(* Logix 5000 project; controller _GigaDiscovery vendor 1 type 14 code 244 rev 35.11; software revision 35.03; part 14 of 23 *)
(* tags used below, declared in another part *)
   Timer : TIMER[60];
   All_Rack_Closed_Mem : BOOL;
   Automatic_E_Stop_Cl_0 : DINT;
   Automatic_E_Stop_Cl_1 : DINT;
   DC_Field_Motor_7 : UDT_CROUT;   // DC Field Motor 7 Gondola Contactor -Q16101E -Q16103E
   DC_Field_Pylon_Motors : UDT_CROUT;   // DC Field Pylon Motors Contactor -Q10101E -Q10103E
   Emergencies_CL0 : DINT[8];
   Emergencies_CL1 : DINT[14];
   FeedBack_Drives_Contactors : BOOL;
   Gondola_Drive_Enable : UDT_CROUT;   // Gondola Drive Ch1-Ch2 Start Enable Contactors -Q16105E -Q16107E
   I_Compressor_Min_Pressure : BOOL;   // Line Pressure Switch - Minimum Pressure -S21504B
   I_EStop_Pb_OCC1 : UDT_DCI_STOP_TEST;   // +OCC E-stop -S30301F
   I_EStop_Pb_OCC2 : UDT_DCI_STOP_TEST;   // +OCC2 E-Stop -S28502F
   I_Gate_ENTER_G01_Closed : UDT_DCM;   // GATE ENTER (G01) -B25204I
   I_Gate_EXIT_G05_Closed : UDT_DCM;   // GATE EXIT (G05) -B25304I
   I_Gate_OPERATOR_Closed : UDT_DCM;   // GATE 4 OPERATOR RFID SENSOR - MOP -B25404J
   I_Gates_Closed : UDT_DCM;   // Gate Closed RFID series -B24802J
   I_OCC1_Stop_Cycle_PB : BOOL;   // Stop Cycle -S30308F
   I_OCC2_ACONFIRM : BOOL;   // OCC2 Allow Main CONFIRM -S28602F
   I_OCC2_Disable : UDT_DCM;   // OCC 2 CONTROL DISABLE Page 310
   I_OCC2_Stop_Cycle_PB : BOOL;   // Stop Cycle -S28606F
   I_OCC_LockOut_Motion : UDT_DCM;   // OCC -Lockout Motion -Q31203E
   I_OCC_Memory_Footpedal : BOOL;
   I_OCC_Operator_Enable_Key : BOOL;   // OCC Console Enabled -S30305F
   I_Operator_Footpedal : BOOL;   // Operator Footpedal -S30901F
   I_Platform_Line_Min_Pressure_Switch : BOOL;   // Platform Line Minimum Pressure Switch -S21511B
   I_Platform_Line_Unlock_Pressure_Switch : BOOL;   // Unlock Platform Line Pressure Switch -S22006B
   I_Platform_Opened : UDT_DCM;   // Platform Opened RFID Series -Q23801J -Q23807J
   I_RESTRAINTS_MainValve_Cosed : BOOL;   // Main Valve Close Limit Switch -B40508I
   I_RESTRAINTS_PressureswitchCompressor : BOOL;   // RESTRAINTS Main Valve Pressure Switch -S40602J
   I_Start_PB : Start_AOI;   // Primary console Strat Push botton Right and Left -S30401F -S30403F
   Mem_All_Rack_Sensor_OFF : BOOL;
   Mem_RESTRAINTS_closed_Correctly : BOOL;
   No_Automatic_E_Stop_Cl_0_Request : BOOL;
   No_Automatic_E_Stop_Cl_1_Request : BOOL;
   No_Emergencies_CL0 : BOOL;
   No_Emergencies_CL1 : BOOL;
   No_Sfty : Std_to_Sfty;
   O_Platform_MainValve : UDT_CROUT;   // Platform main valve B21902I
   O_RESTRAINTS_MainValve : UDT_CROUT;   // Main Valve -B40501I
   Pb_Platform_Stop : BOOL;   // Platform Stop Command -S30608F
   Platform_Open_Cycle : Sequencer;
   Platform_Open_Permissive : Permissive;
   PltaformOpeneded_CycleComplete : BOOL;   // Rilevazione Piattaforme aperte con ciclo Completato
   Power_On_Delay : BOOL;
   ProofTest_Req : BOOL;
   Pylon_Contactor_OFF : BOOL;
   Pylon_Start_Drive_1_2 : UDT_CROUT;   // Pylon Start Drive 1 - 2 Contactors -Q9002H -Q9004H -Q10202G
   Pylon_Start_Drive_3_4 : UDT_CROUT;   // Pylon Start Drive 3 - 4 Contactors -Q9005H -Q9007H -Q12202G
   Pylon_Start_Drive_5_6 : UDT_CROUT;   // Pylon Start Drive 5 - 6 Contactors -Q9009E -Q9011E4 -Q14202G -Q14202G
   Pylon_Stopped_At_Home : BOOL;   // 5s
   Reset_Pulse : BOOL;
   RESTRAINTS_ChA_Open_Memory : BOOL;
   RESTRAINTS_ChB_Open_Memory : BOOL;
   RESTRAINTS_Closed : BOOL;   // All RESTRAINTS Closed
   RESTRAINTS_Rack_Sector_ON : BOOL;
   RESTRAINTS_Sector_Enable_OFF : BOOL;   // ALL RESTRAINTS rack commands OFF
   RESTRAINTS_Unlock_Valve_Pressure : BOOL;
   Start_Permissive : Permissive;
   Start_Permissive2 : Permissive;
   Start_Platform_AutoCycle_Pylon : BOOL;
   Start_Stop_Cycle : Sequencer;
   Start_TOF : TIMER;
   Valve_Proof_Test_Ok : BOOL;
(* S_Alarms, continued *)

ROUTINE _08_Gates   (* ladder *)
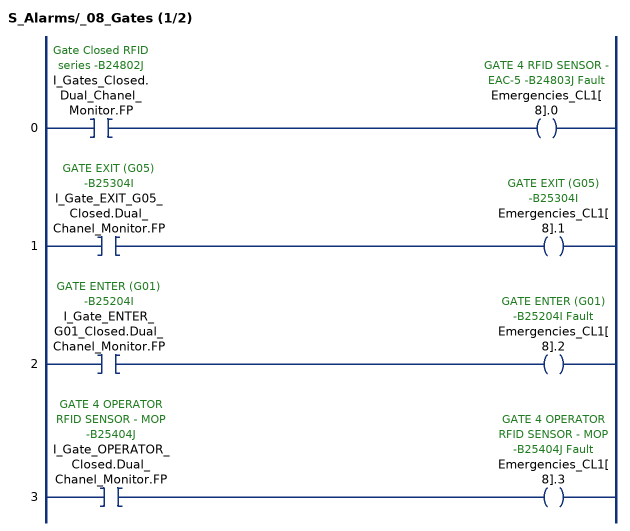
   0: XIC(I_Gates_Closed.Dual_Chanel_Monitor.FP)OTE(Emergencies_CL1[8].0);
   1: XIC(I_Gate_EXIT_G05_Closed.Dual_Chanel_Monitor.FP)OTE(Emergencies_CL1[8].1);
   2: XIC(I_Gate_ENTER_G01_Closed.Dual_Chanel_Monitor.FP)OTE(Emergencies_CL1[8].2);
   3: XIC(I_Gate_OPERATOR_Closed.Dual_Chanel_Monitor.FP)OTE(Emergencies_CL1[8].3);
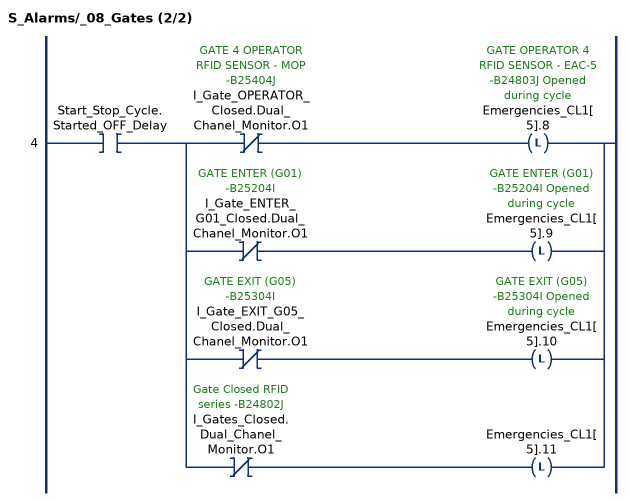
   4: XIC(Start_Stop_Cycle.Started_OFF_Delay)[XIO(I_Gate_OPERATOR_Closed.Dual_Chanel_Monitor.O1) OTL(Emergencies_CL1[5].8) ,XIO(I_Gate_ENTER_G01_Closed.Dual_Chanel_Monitor.O1) OTL(Emergencies_CL1[5].9) ,XIO(I_Gate_EXIT_G05_Closed.Dual_Chanel_Monitor.O1) OTL(Emergencies_CL1[5].10) ,XIO(I_Gates_Closed.Dual_Chanel_Monitor.O1) OTL(Emergencies_CL1[5].11) ];
END_ROUTINE

ROUTINE Main   (* ladder *)
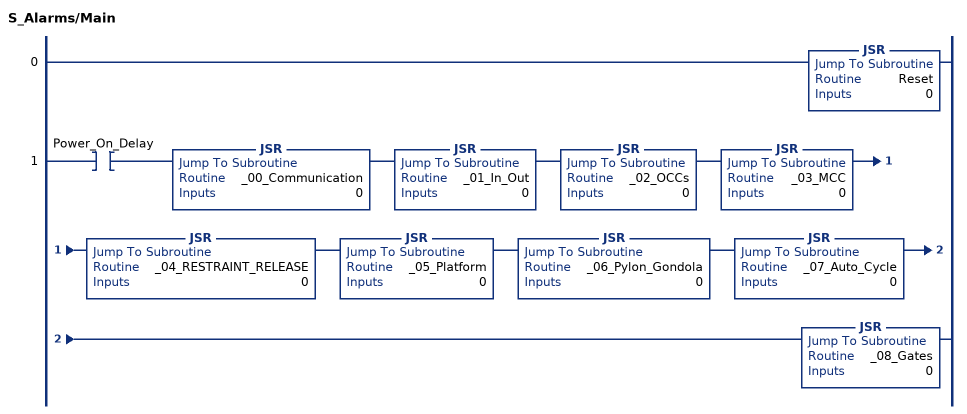
   0: JSR(Reset,0);
   1: XIC(Power_On_Delay)JSR(_00_Communication,0)JSR(_01_In_Out,0)JSR(_02_OCCs,0)JSR(_03_MCC,0)JSR(_04_RESTRAINT_RELEASE,0)JSR(_05_Platform,0)JSR(_06_Pylon_Gondola,0)JSR(_07_Auto_Cycle,0)JSR(_08_Gates,0);
END_ROUTINE

ROUTINE Reset   (* ladder *)
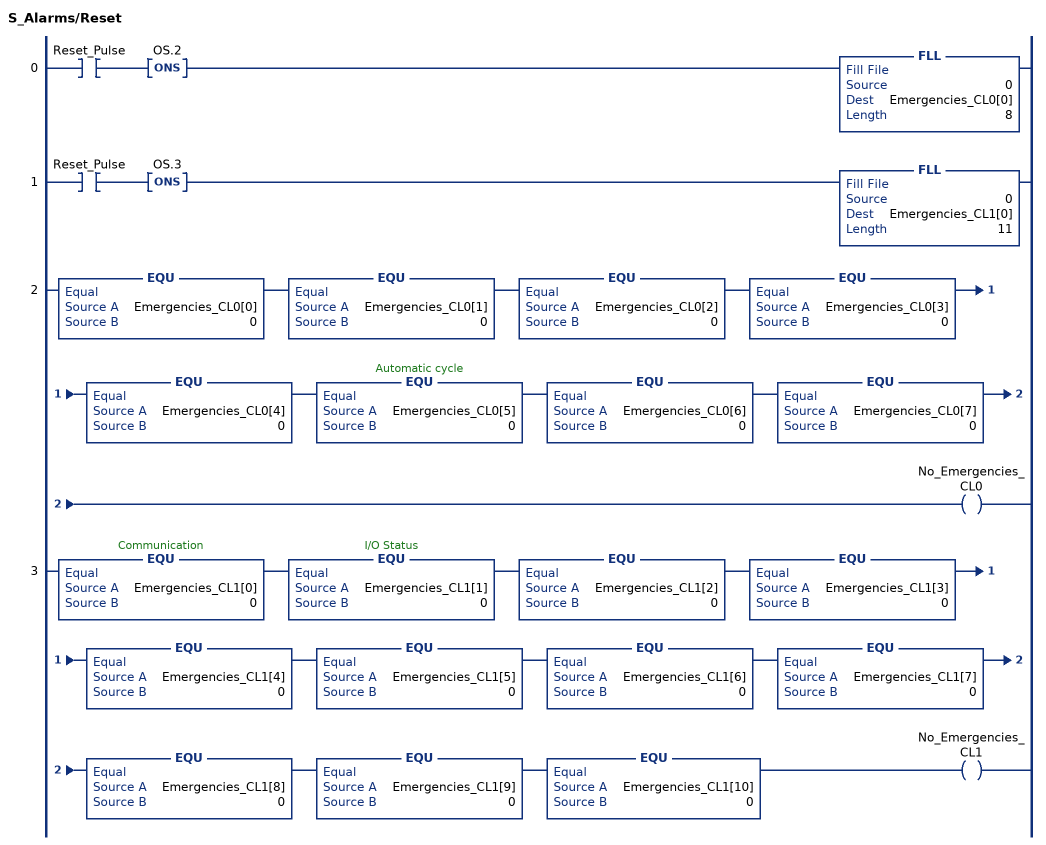
   0: XIC(Reset_Pulse)ONS(OS.2)FLL(0,Emergencies_CL0[0],8);
   1: XIC(Reset_Pulse)ONS(OS.3)FLL(0,Emergencies_CL1[0],11);
   2: EQU(Emergencies_CL0[0],0)EQU(Emergencies_CL0[1],0)EQU(Emergencies_CL0[2],0)EQU(Emergencies_CL0[3],0)EQU(Emergencies_CL0[4],0)EQU(Emergencies_CL0[5],0)EQU(Emergencies_CL0[6],0)EQU(Emergencies_CL0[7],0)OTE(No_Emergencies_CL0);
   3: EQU(Emergencies_CL1[0],0)EQU(Emergencies_CL1[1],0)EQU(Emergencies_CL1[2],0)EQU(Emergencies_CL1[3],0)EQU(Emergencies_CL1[4],0)EQU(Emergencies_CL1[5],0)EQU(Emergencies_CL1[6],0)EQU(Emergencies_CL1[7],0)EQU(Emergencies_CL1[8],0)EQU(Emergencies_CL1[9],0)EQU(Emergencies_CL1[10],0)OTE(No_Emergencies_CL1);
END_ROUTINE
END_PROGRAM

PROGRAM S_Cycles   (* main routine Main, safety *)
VAR
   Brake_Delay : TIMER := (PRE := 10000, ACC := 10000, EN := 1, DN := 1);
   Cycle_AOI : Sequencer_AOI;
   Os : DINT := 4227078;
   Power_On_Delay_Timer : TIMER := (PRE := 80000, ACC := 80000, EN := 1, DN := 1);
   Start_Permissive2_Edge_Fails : DINT := -3;
   Start_Permissive_FailEdge : DINT := -32769;
   Timer_Loc : TIMER[50] := ([0].PRE := 100000, [0].EN := 1, [0].DN := 1, [1].PRE := 500, [2].PRE := 60000, [3].PRE := 5000, [4].PRE := 2100, [4].ACC := 2120, [4].EN := 1, [4].DN := 1, [5].PRE := 10000, [5].ACC := 10000);
END_VAR

ROUTINE _01_Emerg   (* ladder *)
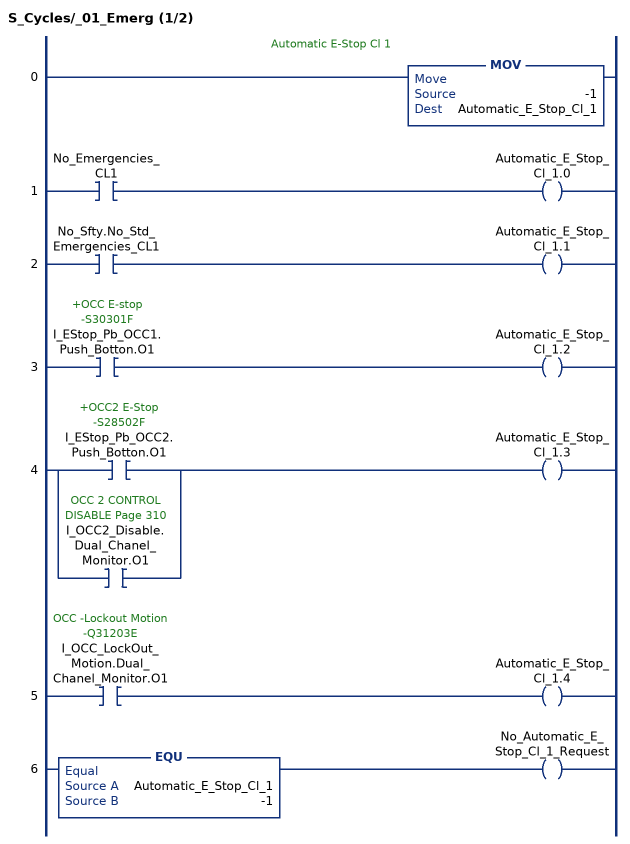
   // Automatic E-Stop Cl 1
   0: MOV(-1,Automatic_E_Stop_Cl_1);
   1: XIC(No_Emergencies_CL1)OTE(Automatic_E_Stop_Cl_1.0);
   2: XIC(No_Sfty.No_Std_Emergencies_CL1)OTE(Automatic_E_Stop_Cl_1.1);
   3: XIC(I_EStop_Pb_OCC1.Push_Botton.O1)OTE(Automatic_E_Stop_Cl_1.2);
   4: [XIC(I_EStop_Pb_OCC2.Push_Botton.O1) ,XIC(I_OCC2_Disable.Dual_Chanel_Monitor.O1) ]OTE(Automatic_E_Stop_Cl_1.3);
   5: XIC(I_OCC_LockOut_Motion.Dual_Chanel_Monitor.O1)OTE(Automatic_E_Stop_Cl_1.4);
   6: EQU(Automatic_E_Stop_Cl_1,-1)OTE(No_Automatic_E_Stop_Cl_1_Request);
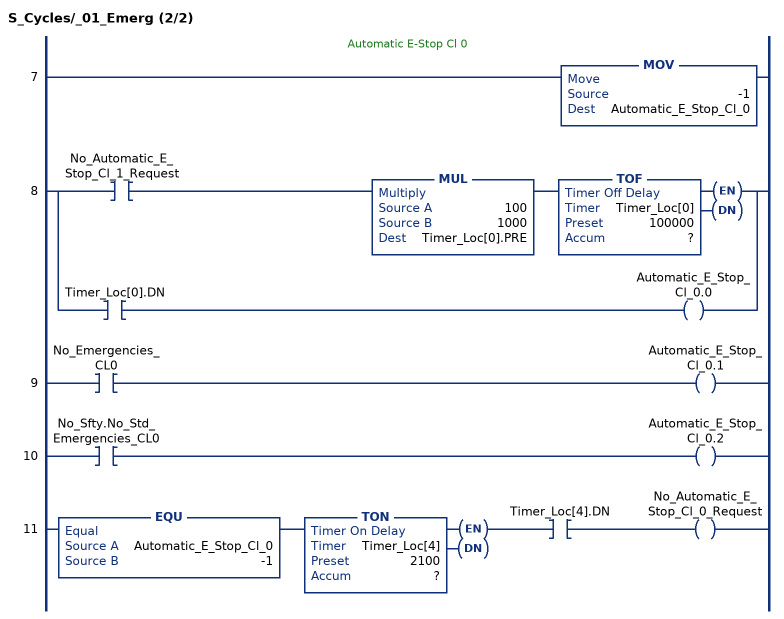
   // Automatic E-Stop Cl 0
   7: MOV(-1,Automatic_E_Stop_Cl_0);
   8: [XIC(No_Automatic_E_Stop_Cl_1_Request) MUL(100,1000,Timer_Loc[0].PRE) TOF(Timer_Loc[0],?,?) ,XIC(Timer_Loc[0].DN) OTE(Automatic_E_Stop_Cl_0.0) ];
   9: XIC(No_Emergencies_CL0)OTE(Automatic_E_Stop_Cl_0.1);
   10: XIC(No_Sfty.No_Std_Emergencies_CL0)OTE(Automatic_E_Stop_Cl_0.2);
   11: EQU(Automatic_E_Stop_Cl_0,-1)TON(Timer_Loc[4],?,?)XIC(Timer_Loc[4].DN)OTE(No_Automatic_E_Stop_Cl_0_Request);
END_ROUTINE

ROUTINE _02_Start_Permissive   (* ladder *)
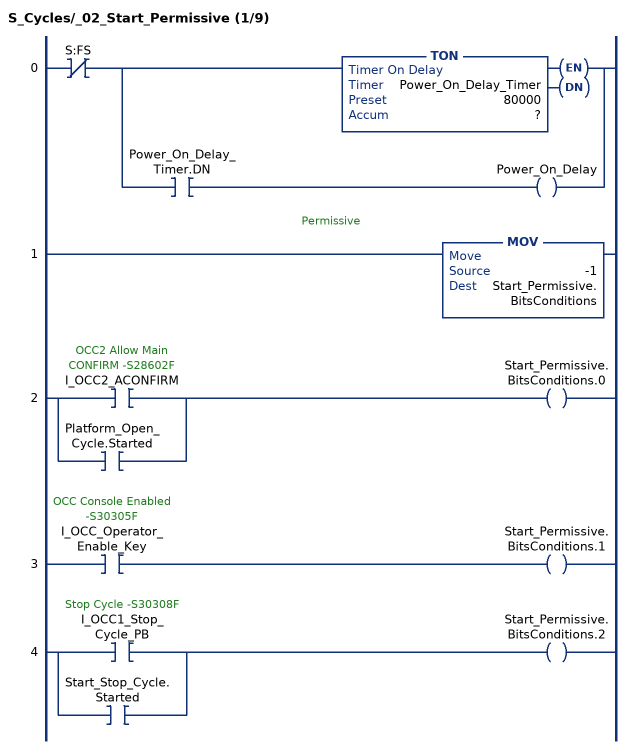
   0: XIO(S:FS)[TON(Power_On_Delay_Timer,?,?) ,XIC(Power_On_Delay_Timer.DN) OTE(Power_On_Delay) ];
   // Permissive
   1: MOV(-1,Start_Permissive.BitsConditions);
   2: [XIC(I_OCC2_ACONFIRM) ,XIC(Platform_Open_Cycle.Started) ]OTE(Start_Permissive.BitsConditions.0);
   3: XIC(I_OCC_Operator_Enable_Key)OTE(Start_Permissive.BitsConditions.1);
   4: [XIC(I_OCC1_Stop_Cycle_PB) ,XIC(Start_Stop_Cycle.Started) ]OTE(Start_Permissive.BitsConditions.2);
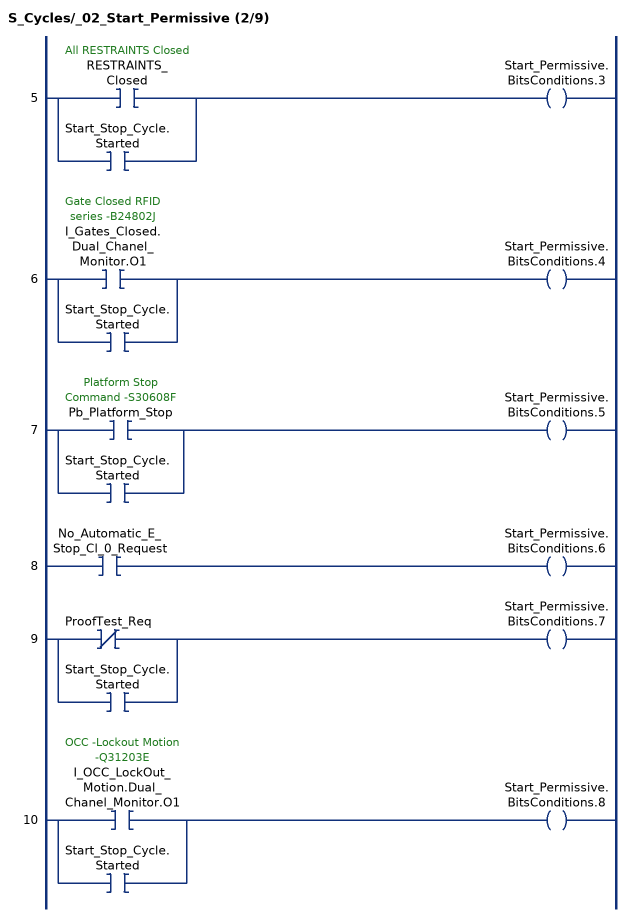
   5: [XIC(RESTRAINTS_Closed) ,XIC(Start_Stop_Cycle.Started) ]OTE(Start_Permissive.BitsConditions.3);
   6: [XIC(I_Gates_Closed.Dual_Chanel_Monitor.O1) ,XIC(Start_Stop_Cycle.Started) ]OTE(Start_Permissive.BitsConditions.4);
   7: [XIC(Pb_Platform_Stop) ,XIC(Start_Stop_Cycle.Started) ]OTE(Start_Permissive.BitsConditions.5);
   8: XIC(No_Automatic_E_Stop_Cl_0_Request)OTE(Start_Permissive.BitsConditions.6);
   9: [XIO(ProofTest_Req) ,XIC(Start_Stop_Cycle.Started) ]OTE(Start_Permissive.BitsConditions.7);
   10: [XIC(I_OCC_LockOut_Motion.Dual_Chanel_Monitor.O1) ,XIC(Start_Stop_Cycle.Started) ]OTE(Start_Permissive.BitsConditions.8);
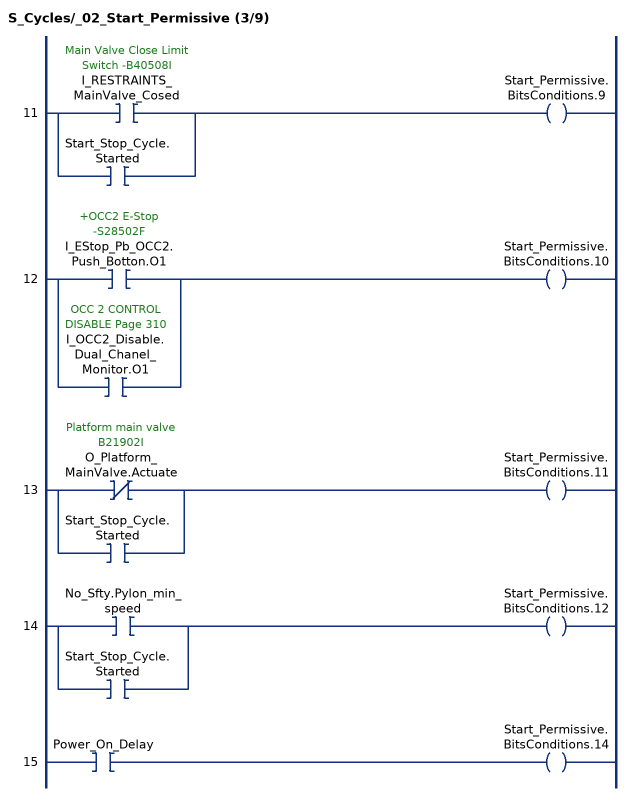
   11: [XIC(I_RESTRAINTS_MainValve_Cosed) ,XIC(Start_Stop_Cycle.Started) ]OTE(Start_Permissive.BitsConditions.9);
   12: [XIC(I_EStop_Pb_OCC2.Push_Botton.O1) ,XIC(I_OCC2_Disable.Dual_Chanel_Monitor.O1) ]OTE(Start_Permissive.BitsConditions.10);
   13: [XIO(O_Platform_MainValve.Actuate) ,XIC(Start_Stop_Cycle.Started) ]OTE(Start_Permissive.BitsConditions.11);
   14: [XIC(No_Sfty.Pylon_min_speed) ,XIC(Start_Stop_Cycle.Started) ]OTE(Start_Permissive.BitsConditions.12);
   15: XIC(Power_On_Delay)OTE(Start_Permissive.BitsConditions.14);
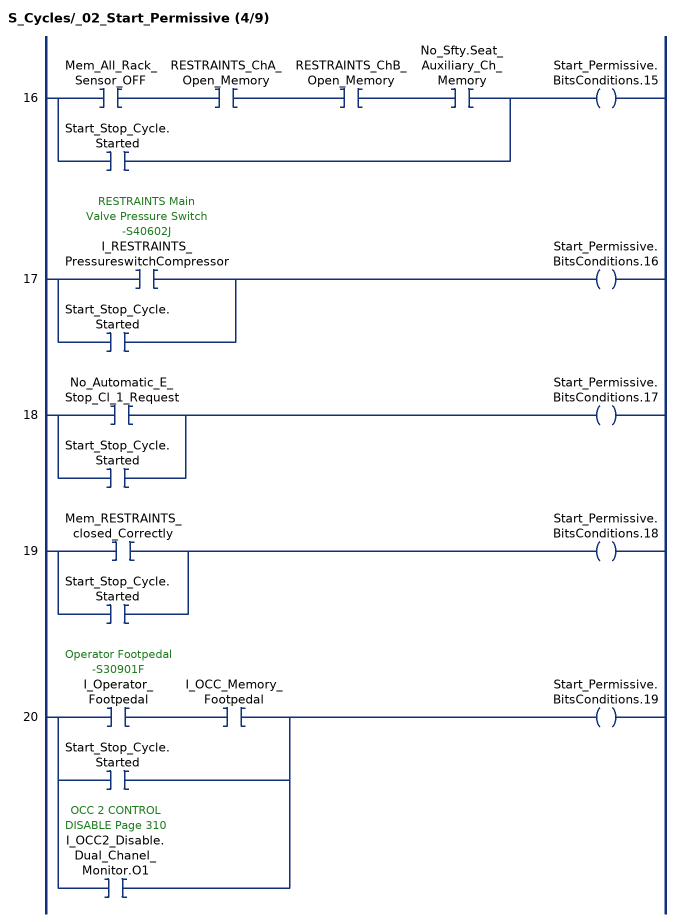
   16: [XIC(Mem_All_Rack_Sensor_OFF) XIC(RESTRAINTS_ChA_Open_Memory) XIC(RESTRAINTS_ChB_Open_Memory) XIC(No_Sfty.Seat_Auxiliary_Ch_Memory) ,XIC(Start_Stop_Cycle.Started) ]OTE(Start_Permissive.BitsConditions.15);
   17: [XIC(I_RESTRAINTS_PressureswitchCompressor) ,XIC(Start_Stop_Cycle.Started) ]OTE(Start_Permissive.BitsConditions.16);
   18: [XIC(No_Automatic_E_Stop_Cl_1_Request) ,XIC(Start_Stop_Cycle.Started) ]OTE(Start_Permissive.BitsConditions.17);
   19: [XIC(Mem_RESTRAINTS_closed_Correctly) ,XIC(Start_Stop_Cycle.Started) ]OTE(Start_Permissive.BitsConditions.18);
   20: [XIC(I_Operator_Footpedal) XIC(I_OCC_Memory_Footpedal) ,XIC(Start_Stop_Cycle.Started) ,XIC(I_OCC2_Disable.Dual_Chanel_Monitor.O1) ]OTE(Start_Permissive.BitsConditions.19);
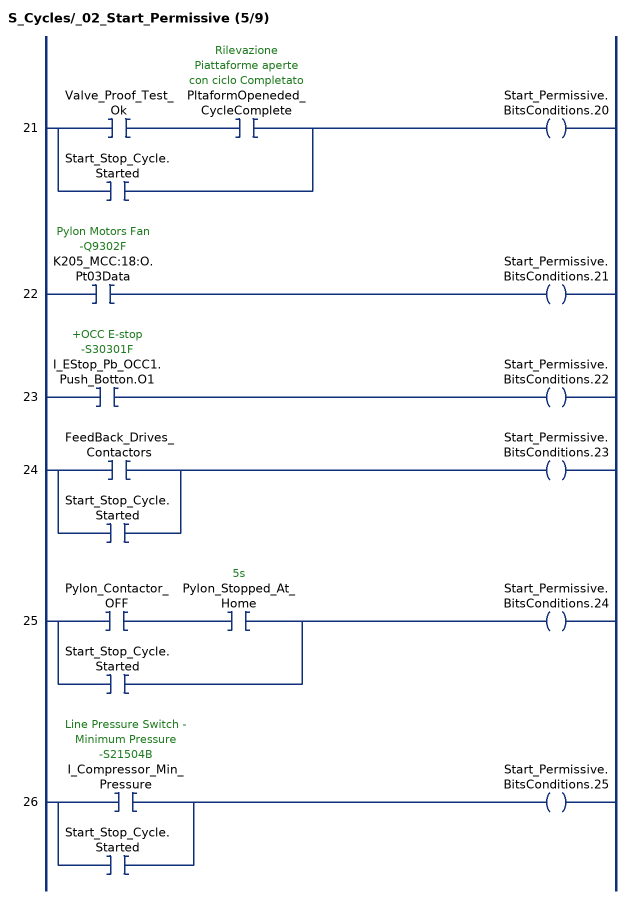
   21: [XIC(Valve_Proof_Test_Ok) XIC(PltaformOpeneded_CycleComplete) ,XIC(Start_Stop_Cycle.Started) ]OTE(Start_Permissive.BitsConditions.20);
   22: XIC(K205_MCC:18:O.Pt03Data)OTE(Start_Permissive.BitsConditions.21);
   23: XIC(I_EStop_Pb_OCC1.Push_Botton.O1)OTE(Start_Permissive.BitsConditions.22);
   24: [XIC(FeedBack_Drives_Contactors) ,XIC(Start_Stop_Cycle.Started) ]OTE(Start_Permissive.BitsConditions.23);
   25: [XIC(Pylon_Contactor_OFF) XIC(Pylon_Stopped_At_Home) ,XIC(Start_Stop_Cycle.Started) ]OTE(Start_Permissive.BitsConditions.24);
   26: [XIC(I_Compressor_Min_Pressure) ,XIC(Start_Stop_Cycle.Started) ]OTE(Start_Permissive.BitsConditions.25);
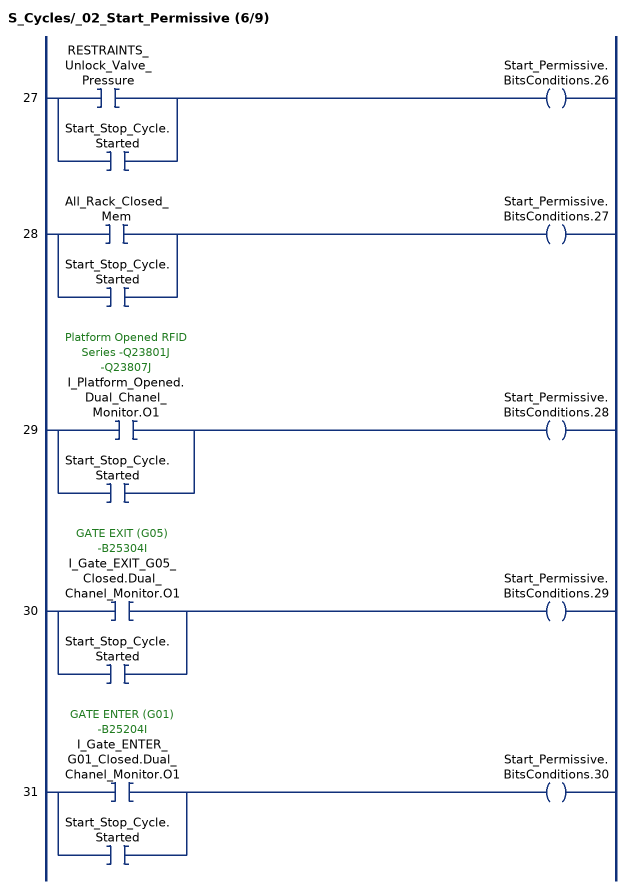
   27: [XIC(RESTRAINTS_Unlock_Valve_Pressure) ,XIC(Start_Stop_Cycle.Started) ]OTE(Start_Permissive.BitsConditions.26);
   28: [XIC(All_Rack_Closed_Mem) ,XIC(Start_Stop_Cycle.Started) ]OTE(Start_Permissive.BitsConditions.27);
   29: [XIC(I_Platform_Opened.Dual_Chanel_Monitor.O1) ,XIC(Start_Stop_Cycle.Started) ]OTE(Start_Permissive.BitsConditions.28);
   30: [XIC(I_Gate_EXIT_G05_Closed.Dual_Chanel_Monitor.O1) ,XIC(Start_Stop_Cycle.Started) ]OTE(Start_Permissive.BitsConditions.29);
   31: [XIC(I_Gate_ENTER_G01_Closed.Dual_Chanel_Monitor.O1) ,XIC(Start_Stop_Cycle.Started) ]OTE(Start_Permissive.BitsConditions.30);
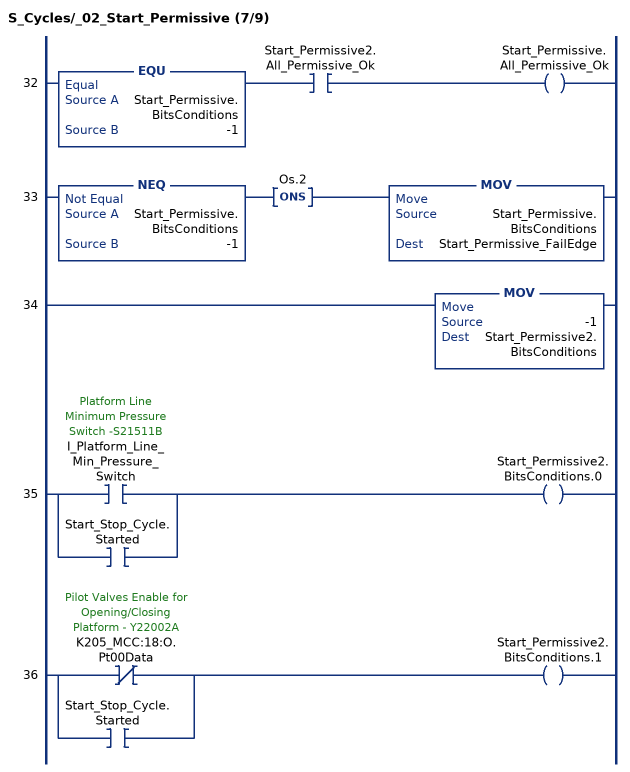
   32: EQU(Start_Permissive.BitsConditions,-1)XIC(Start_Permissive2.All_Permissive_Ok)OTE(Start_Permissive.All_Permissive_Ok);
   33: NEQ(Start_Permissive.BitsConditions,-1)ONS(Os.2)MOV(Start_Permissive.BitsConditions,Start_Permissive_FailEdge);
   34: MOV(-1,Start_Permissive2.BitsConditions);
   35: [XIC(I_Platform_Line_Min_Pressure_Switch) ,XIC(Start_Stop_Cycle.Started) ]OTE(Start_Permissive2.BitsConditions.0);
   36: [XIO(K205_MCC:18:O.Pt00Data) ,XIC(Start_Stop_Cycle.Started) ]OTE(Start_Permissive2.BitsConditions.1);
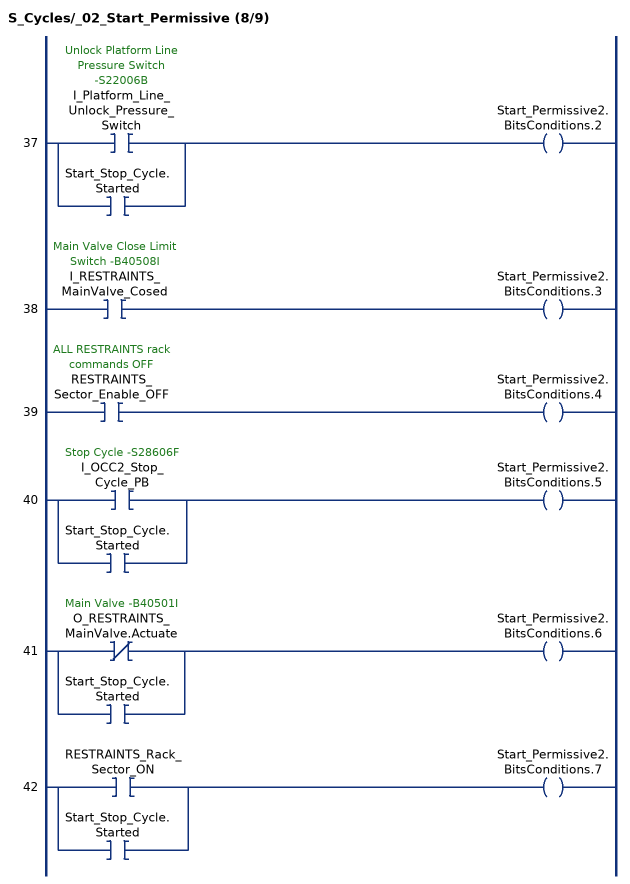
   37: [XIC(I_Platform_Line_Unlock_Pressure_Switch) ,XIC(Start_Stop_Cycle.Started) ]OTE(Start_Permissive2.BitsConditions.2);
   38: XIC(I_RESTRAINTS_MainValve_Cosed)OTE(Start_Permissive2.BitsConditions.3);
   39: XIC(RESTRAINTS_Sector_Enable_OFF)OTE(Start_Permissive2.BitsConditions.4);
   40: [XIC(I_OCC2_Stop_Cycle_PB) ,XIC(Start_Stop_Cycle.Started) ]OTE(Start_Permissive2.BitsConditions.5);
   41: [XIO(O_RESTRAINTS_MainValve.Actuate) ,XIC(Start_Stop_Cycle.Started) ]OTE(Start_Permissive2.BitsConditions.6);
   42: [XIC(RESTRAINTS_Rack_Sector_ON) ,XIC(Start_Stop_Cycle.Started) ]OTE(Start_Permissive2.BitsConditions.7);
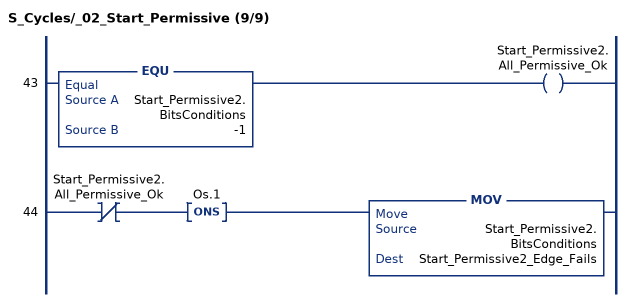
   43: EQU(Start_Permissive2.BitsConditions,-1)OTE(Start_Permissive2.All_Permissive_Ok);
   44: XIO(Start_Permissive2.All_Permissive_Ok)ONS(Os.1)MOV(Start_Permissive2.BitsConditions,Start_Permissive2_Edge_Fails);
END_ROUTINE

ROUTINE _03_Start_Stop_Cycle   (* ladder *)
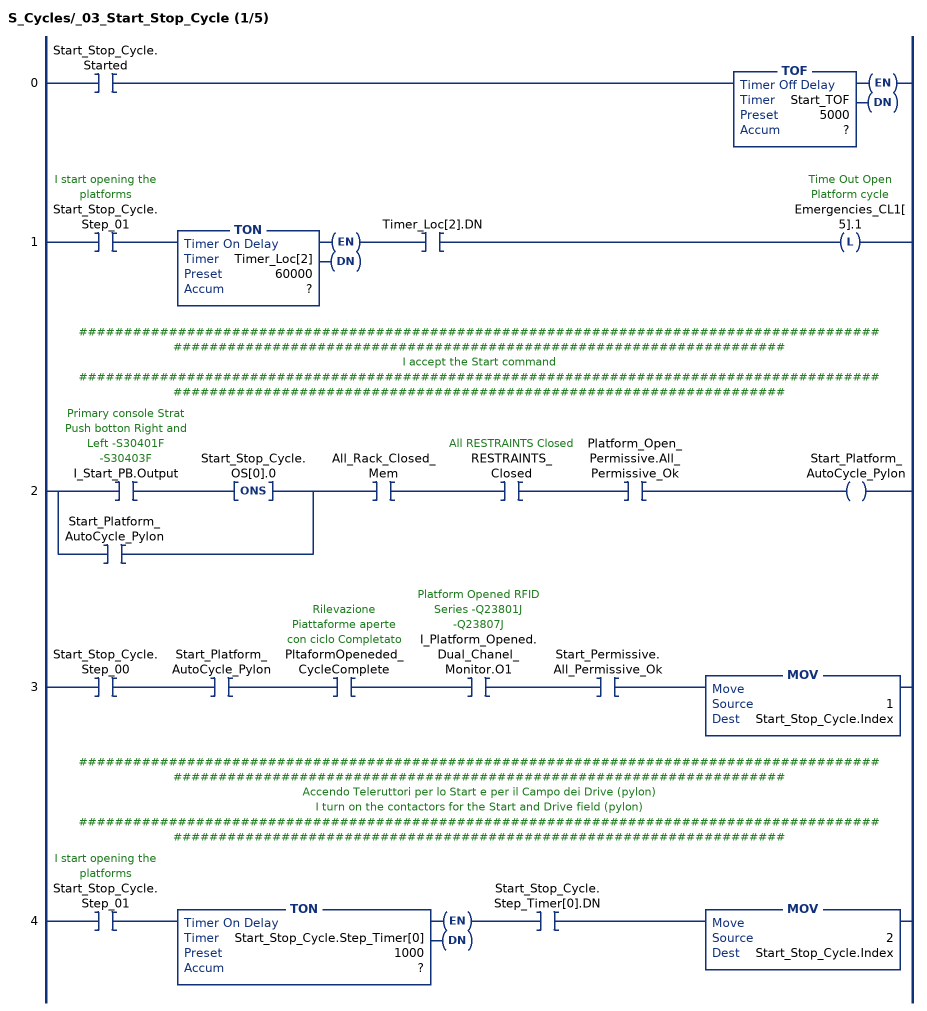
   0: XIC(Start_Stop_Cycle.Started)TOF(Start_TOF,?,?);
   1: XIC(Start_Stop_Cycle.Step_01)TON(Timer_Loc[2],?,?)XIC(Timer_Loc[2].DN)OTL(Emergencies_CL1[5].1);
   // #############################################################################################################################################################
   // I accept the Start command
   // #############################################################################################################################################################
   2: [XIC(I_Start_PB.Output) ONS(Start_Stop_Cycle.OS[0].0) ,XIC(Start_Platform_AutoCycle_Pylon) ]XIC(All_Rack_Closed_Mem)XIC(RESTRAINTS_Closed)XIC(Platform_Open_Permissive.All_Permissive_Ok)OTE(Start_Platform_AutoCycle_Pylon);
   3: XIC(Start_Stop_Cycle.Step_00)XIC(Start_Platform_AutoCycle_Pylon)XIC(PltaformOpeneded_CycleComplete)XIC(I_Platform_Opened.Dual_Chanel_Monitor.O1)XIC(Start_Permissive.All_Permissive_Ok)MOV(1,Start_Stop_Cycle.Index);
   // #############################################################################################################################################################
   // Accendo Teleruttori per lo Start e per il Campo dei Drive (pylon)
   // I turn on the contactors for the Start and Drive field (pylon)
   // #############################################################################################################################################################
   4: XIC(Start_Stop_Cycle.Step_01)TON(Start_Stop_Cycle.Step_Timer[0],?,?)XIC(Start_Stop_Cycle.Step_Timer[0].DN)MOV(2,Start_Stop_Cycle.Index);
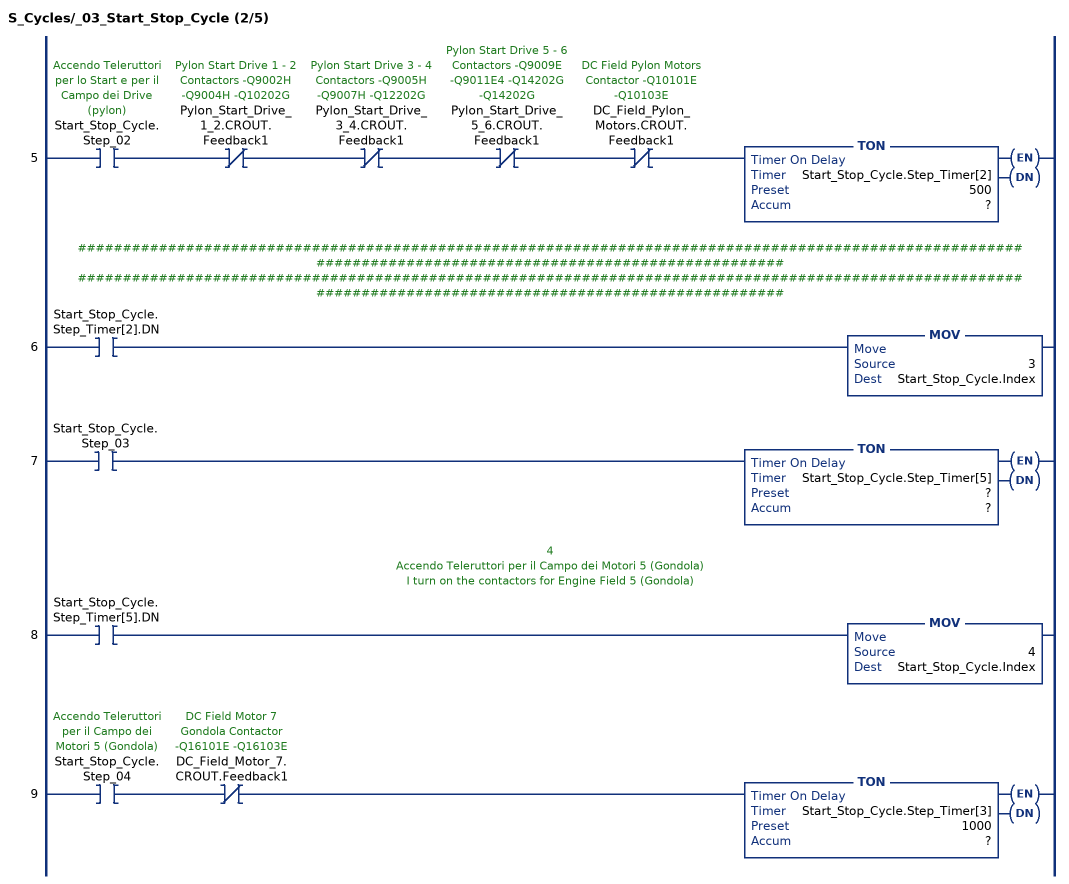
   5: XIC(Start_Stop_Cycle.Step_02)XIO(Pylon_Start_Drive_1_2.CROUT.Feedback1)XIO(Pylon_Start_Drive_3_4.CROUT.Feedback1)XIO(Pylon_Start_Drive_5_6.CROUT.Feedback1)XIO(DC_Field_Pylon_Motors.CROUT.Feedback1)TON(Start_Stop_Cycle.Step_Timer[2],?,?);
   // #############################################################################################################################################################
   // #############################################################################################################################################################
   6: XIC(Start_Stop_Cycle.Step_Timer[2].DN)MOV(3,Start_Stop_Cycle.Index);
   7: XIC(Start_Stop_Cycle.Step_03)TON(Start_Stop_Cycle.Step_Timer[5],?,?);
   // 4
   // Accendo Teleruttori per il Campo dei Motori 5 (Gondola)
   // I turn on the contactors for Engine Field 5 (Gondola)
   8: XIC(Start_Stop_Cycle.Step_Timer[5].DN)MOV(4,Start_Stop_Cycle.Index);
   9: XIC(Start_Stop_Cycle.Step_04)XIO(DC_Field_Motor_7.CROUT.Feedback1)TON(Start_Stop_Cycle.Step_Timer[3],?,?);
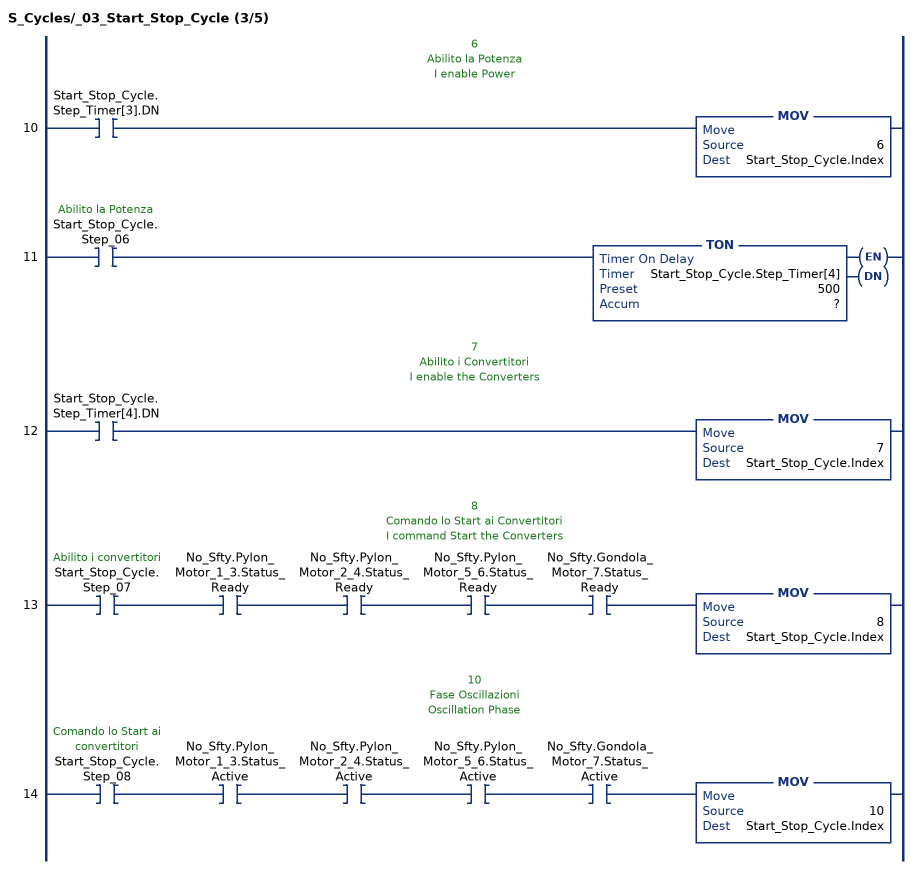
   // 6
   // Abilito la Potenza
   // I enable Power
   10: XIC(Start_Stop_Cycle.Step_Timer[3].DN)MOV(6,Start_Stop_Cycle.Index);
   11: XIC(Start_Stop_Cycle.Step_06)TON(Start_Stop_Cycle.Step_Timer[4],?,?);
   // 7
   // Abilito i Convertitori
   // I enable the Converters
   12: XIC(Start_Stop_Cycle.Step_Timer[4].DN)MOV(7,Start_Stop_Cycle.Index);
   // 8
   // Comando lo Start ai Convertitori
   // I command Start the Converters
   13: XIC(Start_Stop_Cycle.Step_07)XIC(No_Sfty.Pylon_Motor_1_3.Status_Ready)XIC(No_Sfty.Pylon_Motor_2_4.Status_Ready)XIC(No_Sfty.Pylon_Motor_5_6.Status_Ready)XIC(No_Sfty.Gondola_Motor_7.Status_Ready)MOV(8,Start_Stop_Cycle.Index);
   // 10
   // Fase Oscillazioni
   // Oscillation Phase
   14: XIC(Start_Stop_Cycle.Step_08)XIC(No_Sfty.Pylon_Motor_1_3.Status_Active)XIC(No_Sfty.Pylon_Motor_2_4.Status_Active)XIC(No_Sfty.Pylon_Motor_5_6.Status_Active)XIC(No_Sfty.Gondola_Motor_7.Status_Active)MOV(10,Start_Stop_Cycle.Index);
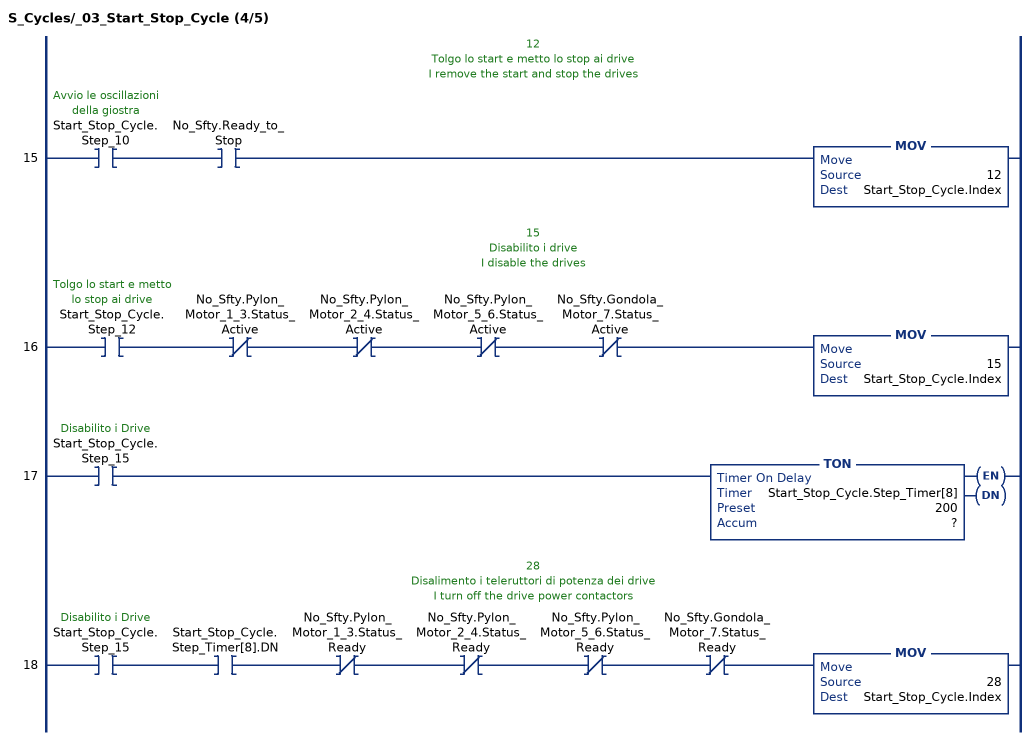
   // 12
   // Tolgo lo start e metto lo stop ai drive
   // I remove the start and stop the drives
   15: XIC(Start_Stop_Cycle.Step_10)XIC(No_Sfty.Ready_to_Stop)MOV(12,Start_Stop_Cycle.Index);
   // 15
   // Disabilito i drive
   // I disable the drives
   16: XIC(Start_Stop_Cycle.Step_12)XIO(No_Sfty.Pylon_Motor_1_3.Status_Active)XIO(No_Sfty.Pylon_Motor_2_4.Status_Active)XIO(No_Sfty.Pylon_Motor_5_6.Status_Active)XIO(No_Sfty.Gondola_Motor_7.Status_Active)MOV(15,Start_Stop_Cycle.Index);
   17: XIC(Start_Stop_Cycle.Step_15)TON(Start_Stop_Cycle.Step_Timer[8],?,?);
   // 28
   // Disalimento i teleruttori di potenza dei drive
   // I turn off the drive power contactors
   18: XIC(Start_Stop_Cycle.Step_15)XIC(Start_Stop_Cycle.Step_Timer[8].DN)XIO(No_Sfty.Pylon_Motor_1_3.Status_Ready)XIO(No_Sfty.Pylon_Motor_2_4.Status_Ready)XIO(No_Sfty.Pylon_Motor_5_6.Status_Ready)XIO(No_Sfty.Gondola_Motor_7.Status_Ready)MOV(28,Start_Stop_Cycle.Index);
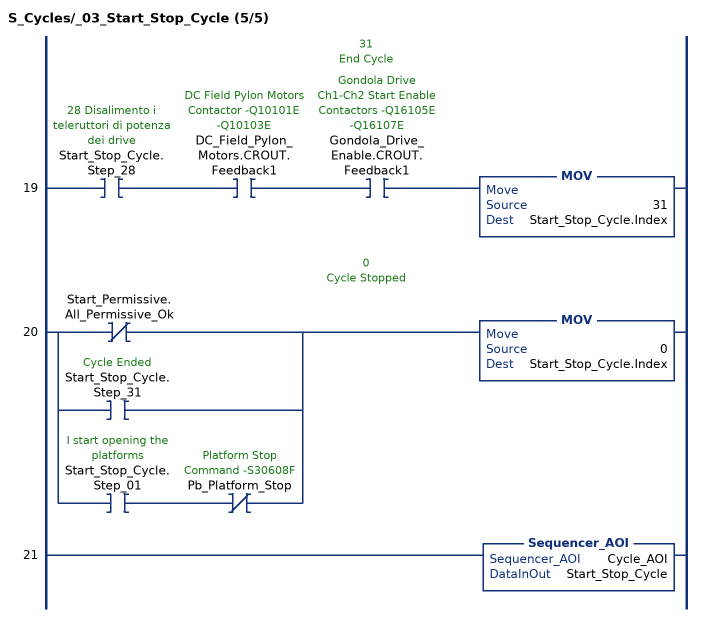
   // 31
   // End Cycle
   19: XIC(Start_Stop_Cycle.Step_28)XIC(DC_Field_Pylon_Motors.CROUT.Feedback1)XIC(Gondola_Drive_Enable.CROUT.Feedback1)MOV(31,Start_Stop_Cycle.Index);
   // 0
   // Cycle Stopped
   20: [XIO(Start_Permissive.All_Permissive_Ok) ,XIC(Start_Stop_Cycle.Step_31) ,XIC(Start_Stop_Cycle.Step_01) XIO(Pb_Platform_Stop) ]MOV(0,Start_Stop_Cycle.Index);
   21: Sequencer_AOI(Cycle_AOI,Start_Stop_Cycle);
END_ROUTINE
